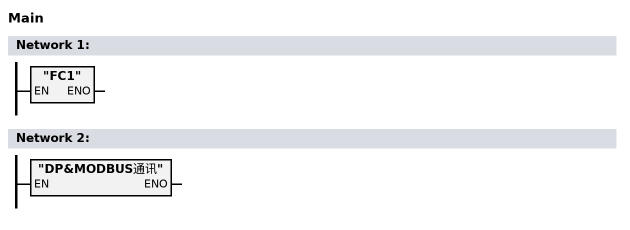
   RUNG wire#powerrail
      "FC1"()
   END_RUNG
   // the same network as SCL:
   "FC1"();
END_REGION

REGION Network 2
   RUNG wire#powerrail
      "DP&MODBUS通讯"()
   END_RUNG
   // the same network as SCL:
   "DP&MODBUS通讯"();
END_REGION
END_ORGANIZATION_BLOCK

// ===== PLC "2#GZY"  CPU 1511-1 PN =====

VAR_GLOBAL   // PLC tag table "默认变量表"
   "Clock_Byte" AT %MB0 : Byte;
   "Clock_10Hz" AT %M0.0 : Bool;
   "Clock_5Hz" AT %M0.1 : Bool;
   "Clock_2.5Hz" AT %M0.2 : Bool;
   "Clock_2Hz" AT %M0.3 : Bool;
   "Clock_1.25Hz" AT %M0.4 : Bool;
   "Clock_1Hz" AT %M0.5 : Bool;
   "Clock_0.625Hz" AT %M0.6 : Bool;
   "Clock_0.5Hz" AT %M0.7 : Bool;
   "2#干燥窑主机远程" AT %I0.0 : Bool;
   "2#干燥窑主机变频备妥" AT %I0.1 : Bool;
   "2#干燥窑主机散热风机运行" AT %I0.2 : Bool;
   "2#干燥窑变频运行" AT %I0.3 : Bool;
   "2#干燥窑变频故障" AT %I0.4 : Bool;
   "2#干燥窑稀油中控" AT %I1.0 : Bool;
   "2#干燥窑稀油1#泵运行" AT %I1.1 : Bool;
   "2#干燥窑稀油2#泵运行" AT %I1.2 : Bool;
   "2#干燥窑稀油油差下限" AT %I1.3 : Bool;
   "2#干燥窑稀油油位上限" AT %I1.4 : Bool;
   "2#干燥窑稀油油位下限" AT %I1.5 : Bool;
   "2#干燥窑稀油1#泵故障" AT %I1.6 : Bool;
   "2#干燥窑稀油2#泵故障" AT %I1.7 : Bool;
   "2#干燥窑挡轮备妥" AT %I2.0 : Bool;
   "2#干燥窑挡轮1#泵运行" AT %I2.1 : Bool;
   "2#干燥窑挡轮2#泵运行" AT %I2.2 : Bool;
   "2#干燥窑挡轮溢流阀运行" AT %I2.3 : Bool;
   "2#干燥窑挡轮行程过低" AT %I2.4 : Bool;
   "2#干燥窑挡轮故障" AT %I2.5 : Bool;
   "I3_0" AT %I3.0 : Bool;
   "I3_1" AT %I3.1 : Bool;
   "I3_2" AT %I3.2 : Bool;
   "湿矿转2#干燥窑皮中控  (3#皮带)" AT %I3.3 : Bool;
   "湿矿转2#干燥窑皮运行  (3#皮带)" AT %I3.4 : Bool;
   "湿矿转2#干燥窑皮故障  (3#皮带)" AT %I3.5 : Bool;
   "I4_0" AT %I4.0 : Bool;
   "I4_1" AT %I4.1 : Bool;
   "I4_2" AT %I4.2 : Bool;
   "I4_3" AT %I4.3 : Bool;
   "I4_4" AT %I4.4 : Bool;
   "I4_5" AT %I4.5 : Bool;
   "I5_0" AT %I5.0 : Bool;
   "I5_1" AT %I5.1 : Bool;
   "I5_2" AT %I5.2 : Bool;
   "I5_3" AT %I5.3 : Bool;
   "I5_4" AT %I5.4 : Bool;
   "I5_5" AT %I5.5 : Bool;
   "定量给煤机中控" AT %I6.3 : Bool;
   "定量给煤机运行" AT %I6.4 : Bool;
   "定量给煤机故障" AT %I6.5 : Bool;
   "定量给煤机流量脉冲" AT %I6.6 : Bool;
   "煤粉仓收尘风机中控" AT %I7.0 : Bool;
   "煤粉仓收尘风机运行" AT %I7.1 : Bool;
   "煤粉仓收尘风机故障" AT %I7.2 : Bool;
   "2#干燥窑一次风机中控" AT %I8.0 : Bool;
   "2#干燥窑一次风机运行" AT %I8.1 : Bool;
   "2#干燥窑一次风机故障" AT %I8.2 : Bool;
   "2#干燥窑二次风机中控" AT %I8.3 : Bool;
   "2#干燥窑二次风机运行" AT %I8.4 : Bool;
   "2#干燥窑二次风机故障" AT %I8.5 : Bool;
   "I9_0" AT %I9.0 : Bool;
   "I9_1" AT %I9.1 : Bool;
   "I9_2" AT %I9.2 : Bool;
   "I9_3" AT %I9.3 : Bool;
   "I9_4" AT %I9.4 : Bool;
   "I9_5" AT %I9.5 : Bool;
   "I10_0" AT %I10.0 : Bool;
   "I10_1" AT %I10.1 : Bool;
   "I10_2" AT %I10.2 : Bool;
   "I10_4" AT %I10.4 : Bool;
   "I10_5" AT %I10.5 : Bool;
   "I10_6" AT %I10.6 : Bool;
   "2#干燥窑转速" AT %IW256 : Int;
   "2#干燥窑电流" AT %IW258 : Int;
   "PIW260" AT %IW260 : Int;
   "2#干燥窑一次风机电流" AT %IW262 : Int;
   "2#干燥窑二次风机频率" AT %IW264 : Int;
   "2#干燥窑二次风机电流" AT %IW266 : Int;
   "PIW268" AT %IW268 : Int;
   "PIW270" AT %IW270 : Int;
   "2#干燥窑窑尾压力" AT %IW272 : Int;
   "PIW274" AT %IW274 : Int;
   "定量给煤机流量" AT %IW276 : Int;
   "烟气管道进口压力" AT %IW278 : Int;
   "2#干燥窑一次风压" AT %IW280 : Int;
   "2#干燥窑二次风压" AT %IW282 : Int;
   "煤粉仓压力" AT %IW284 : Int;
   "混合室压力" AT %IW286 : Int;
   "煤粉仓温度1(PT100)" AT %IW288 : Int;
   "煤粉仓温度2(PT100)" AT %IW290 : Int;
   "煤粉仓温度3(PT100)" AT %IW292 : Int;
   "煤粉仓温度4(PT100)" AT %IW294 : Int;
   "窑尾温度 K偶" AT %IW296 : Int;
   "烟气管道进口温度 K偶" AT %IW298 : Int;
   "燃烧室温度 4~20mA" AT %IW300 : Int;
   "混合室温度 4~20mA" AT %IW302 : Int;
   "2#窑A档轴温1" AT %ID320 : Real;
   "2#窑A档油温1" AT %ID324 : Real;
   "2#窑A档轴温2" AT %ID328 : Real;
   "2#窑A档油温2" AT %ID332 : Real;
   "2#窑A档轴温3" AT %ID336 : Real;
   "2#窑A档油温3" AT %ID340 : Real;
   "2#窑A档轴温4" AT %ID344 : Real;
   "2#窑A档油温4" AT %ID348 : Real;
   "2#窑B档轴温1" AT %ID352 : Real;
   "2#窑B档油温1" AT %ID356 : Real;
   "2#窑B档轴温2" AT %ID360 : Real;
   "2#窑B档油温2" AT %ID364 : Real;
   "2#窑B档轴温3" AT %ID368 : Real;
   "2#窑B档油温3" AT %ID372 : Real;
   "2#窑B档轴温4" AT %ID376 : Real;
   "2#窑B档油温4" AT %ID380 : Real;
   "2#窑主电机A相绕组温度" AT %ID384 : Real;
   "干燥窑主传动合闸" AT %Q0.0 : Bool;
   "干燥窑主传动分闸" AT %Q0.1 : Bool;
   "干燥窑主传动变频启动" AT %Q0.2 : Bool;
   "干燥窑主传稀油站启动" AT %Q0.3 : Bool;
   "湿矿转2#干燥窑皮带启动  (3#皮带)" AT %Q0.4 : Bool;
   "Q0_5" AT %Q0.5 : Bool;
   "Q0_6" AT %Q0.6 : Bool;
   "Q0_7" AT %Q0.7 : Bool;
   "Q1_0" AT %Q1.0 : Bool;
   "定量给煤机启动" AT %Q1.2 : Bool;
   "煤粉仓收尘风机启动" AT %Q1.3 : Bool;
   "Q1_4" AT %Q1.4 : Bool;
   "Q1_5" AT %Q1.5 : Bool;
   "干燥窑挡轮油站启动" AT %Q1.6 : Bool;
   "2#干燥窑一次风机启动" AT %Q2.0 : Bool;
   "2#干燥窑二次风机启动" AT %Q2.1 : Bool;
   "Q2_2" AT %Q2.2 : Bool;
   "Q2_3" AT %Q2.3 : Bool;
   "Tag_8" AT %QB4 : Byte;
   "2#干燥窑转速给定" AT %QW256 : Int;
   "定量给煤机流量给定" AT %QW258 : Int;
   "PQW264" AT %QW264 : Int;
   "2#干燥窑二次风机频率给定" AT %QW266 : Int;
   "PQW268" AT %QW268 : Int;
   "PQW270" AT %QW270 : Int;
   "Tag_1" AT %MW4 : Word;
   "Tag_2" AT %M400.0 : Bool;
   "连锁解锁" AT %M400.2 : Bool;
   "干燥窑连锁信号" AT %M400.3 : Bool;
   "Tag_4" AT %M400.5 : Bool;
   "Tag_5" AT %MW410 : Word;
   "Tag_6" AT %MW412 : Word;
   "稀油站油压长时间低" AT %T6 : Timer;
   "稀油站启动10S" AT %T7 : Timer;
   "稀油站油差下限时间" AT %T8 : Timer;
   "Tag_3" AT %C1 : Counter;
   "Tag_7" AT %C2 : Counter;
   "2#干燥窑断路器合闸" AT %I0.5 : Bool;
   "2#干燥窑断路器分闸" AT %I0.6 : Bool;
   "2#干燥窑进料口压力" AT %IW304 : Int;
   "Tag_31" AT %T1 : Timer;
   "Tag_33" AT %T2 : Timer;
   "Q1_1" AT %Q1.1 : Bool;
   "System_Byte" AT %MB1 : Byte;
   "FirstScan" AT %M1.0 : Bool;
   "DiagStatusUpdate" AT %M1.1 : Bool;
   "AlwaysTRUE" AT %M1.2 : Bool;
   "AlwaysFALSE" AT %M1.3 : Bool;
   "2#窑主电机B相绕组温度" AT %ID388 : Real;
   "2#窑主电机C相绕组温度" AT %ID392 : Real;
   "2#窑主电机前轴承温度" AT %ID396 : Real;
   "2#窑主电机后轴承温度" AT %ID400 : Real;
   "I0_7" AT %I0.7 : Bool;
   "I2_6" AT %I2.6 : Bool;
   "I2_7" AT %I2.7 : Bool;
   "I3_6" AT %I3.6 : Bool;
   "I3_7" AT %I3.7 : Bool;
   "I4_6" AT %I4.6 : Bool;
   "I4_7" AT %I4.7 : Bool;
   "I5_6" AT %I5.6 : Bool;
   "I5_7" AT %I5.7 : Bool;
   "I6_0" AT %I6.0 : Bool;
   "I6_1" AT %I6.1 : Bool;
   "I6_2" AT %I6.2 : Bool;
   "I6_7" AT %I6.7 : Bool;
   "I7_3" AT %I7.3 : Bool;
   "I7_4" AT %I7.4 : Bool;
   "I7_5" AT %I7.5 : Bool;
   "I7_6" AT %I7.6 : Bool;
   "I7_7" AT %I7.7 : Bool;
   "I8_6" AT %I8.6 : Bool;
   "I8_7" AT %I8.7 : Bool;
   "I9_6" AT %I9.6 : Bool;
   "I9_7" AT %I9.7 : Bool;
   "I10_3" AT %I10.3 : Bool;
   "I10_7" AT %I10.7 : Bool;
   "I11_0" AT %I11.0 : Bool;
   "I11_1" AT %I11.1 : Bool;
   "I11_2" AT %I11.2 : Bool;
   "I11_3" AT %I11.3 : Bool;
   "I11_4" AT %I11.4 : Bool;
   "I11_5" AT %I11.5 : Bool;
   "I11_6" AT %I11.6 : Bool;
   "I11_7" AT %I11.7 : Bool;
   "Q1_7" AT %Q1.7 : Bool;
   "Q2_4" AT %Q2.4 : Bool;
   "Q2_5" AT %Q2.5 : Bool;
   "Q2_6" AT %Q2.6 : Bool;
   "Q2_7" AT %Q2.7 : Bool;
   "Q3_0" AT %Q3.0 : Bool;
   "Q3_1" AT %Q3.1 : Bool;
   "Q3_2" AT %Q3.2 : Bool;
   "Q3_3" AT %Q3.3 : Bool;
   "Q3_4" AT %Q3.4 : Bool;
   "Q3_5" AT %Q3.5 : Bool;
   "Q3_6" AT %Q3.6 : Bool;
   "Q3_7" AT %Q3.7 : Bool;
   "2#给煤机出料口负压" AT %IW306 : Int;
   "PIW308" AT %IW308 : Int;
   "PIW310" AT %IW310 : Int;
   "PIW312" AT %IW312 : Int;
   "PIW314" AT %IW314 : Int;
   "PIW316" AT %IW316 : Int;
   "PIW318" AT %IW318 : Int;
   "PQW260" AT %QW260 : Int;
   "PQW262" AT %QW262 : Int;
   "2#干燥窑煤粉仓称重" AT %ID440 : Real;
   "Tag_9" AT %T10 : Timer;
END_VAR

DATA_BLOCK "驱动"   // DB1
{ S7_Optimized_Access := 'FALSE' }
VERSION : 0.1
   VAR
      "2#二次风机启动" : Bool;
      "2#二次风机停止" : Bool;
      "2#干燥窑主机合闸" : Bool;
      "2#干燥窑主机分闸" : Bool;
      STAT4 : Bool;
      STAT5 : Bool;
      "2#干燥窑主机启动" : Bool;
      "2#干燥窑主机停止" : Bool;
      STAT8 : Bool;
      STAT9 : Bool;
      STAT10 : Bool;
      STAT11 : Bool;
      "gzy进窑2#皮带启动3#皮带" : Bool;
      "gzy进窑2#皮带停止3#皮带" : Bool;
      STAT14 : Bool;
      STAT15 : Bool;
      STAT16 : Bool;
      STAT17 : Bool;
      STAT18 : Bool;
      STAT19 : Bool;
      STAT20 : Bool;
      STAT21 : Bool;
      STAT22 : Bool;
      STAT23 : Bool;
      STAT24 : Bool;
      STAT25 : Bool;
      STAT26 : Bool;
      STAT27 : Bool;
      "2#一次风机启动" : Bool;
      "2#一次风机停止" : Bool;
      STAT30 : Bool;
      STAT31 : Bool;
      STAT32 : Bool;
      STAT33 : Bool;
      STAT34 : Bool;
      STAT35 : Bool;
      STAT36 : Bool;
      STAT37 : Bool;
      STAT38 : Bool;
      STAT39 : Bool;
      "2#干燥窑煤粉收尘风机启动" : Bool;
      "2#干燥窑煤粉收尘风机停止" : Bool;
      "2#干燥窑锁风给煤机启动" : Bool;
      "2#干燥窑锁风给煤机停止" : Bool;
      "2#干燥窑锁风给煤机分割轮启动" : Bool;
      "2#干燥窑锁风给煤机分割轮停止" : Bool;
      STAT46 : Bool;
      STAT47 : Bool;
      STAT48 : Bool;
      STAT49 : Bool;
      STAT50 : Bool;
      STAT51 : Bool;
      STAT52 : Bool;
      STAT53 : Bool;
      STAT54 : Bool;
      STAT55 : Bool;
      STAT56 : Bool;
      "2#干燥窑联锁解锁" : Bool;
      STAT58 : Bool;
      STAT59 : Bool;
      STAT60 : Bool;
      "2#干燥窑定量给煤机班累计清零" : Bool;
      "2#干燥窑定量给煤机日累计清零" : Bool;
      "2#干燥窑定量给煤机总累计清零" : Bool;
      STAT64 : Bool;
      STAT65 : Bool;
      "2#干燥窑稀油站启动" : Bool;
      "2#干燥窑稀油站停止" : Bool;
      "2#干燥窑挡轮油站启动" : Bool;
      "2#干燥窑挡轮油站停止" : Bool;
      STAT66 : Bool;
      STAT67 : Bool;
   END_VAR
BEGIN
END_DATA_BLOCK

DATA_BLOCK "模拟量"   // DB2
{ S7_Optimized_Access := 'FALSE' }
VERSION : 0.1
   VAR
      STAT0 : Int;
      STAT1 : Int;
      STAT2 : Int;
      STAT3 : Int;
      STAT4 : Int;
      STAT5 : Int;
      STAT6 : Int;
      STAT7 : Int;
      STAT8 : Int;
      STAT9 : Real;
      STAT10 : Real;
      STAT11 : Real;
      STAT12 : Real;
      STAT13 : Real;
      STAT14 : Real;
      STAT15 : Real;
      STAT16 : Real;
      STAT17 : Real;
      STAT18 : Real;
      STAT19 : Real;
      STAT20 : Real;
      STAT21 : Real;
      STAT22 : Real;
      STAT23 : Real;
      STAT24 : Real;
      STAT25 : Real;
      STAT26 : Real;
      STAT27 : Real;
      STAT28 : Real;
      STAT29 : Real;
      STAT30 : Real;
      STAT31 : Real;
      STAT32 : Real;
      STAT33 : Real;
      STAT34 : Real;
      STAT35 : Real;
      STAT36 : Real;
      STAT37 : Real;
      STAT38 : Real;
      STAT39 : Real;
      STAT40 : Real;
      STAT41 : Real;
      STAT42 : Real;
      STAT43 : Real;
      STAT44 : Real;
      STAT45 : Real;
      STAT46 : Real;
      STAT47 : Real;
      STAT48 : Real;
      STAT49 : Real;
      STAT50 : Real;
      STAT51 : Real;
      STAT52 : Real;
      STAT53 : Real;
      STAT54 : Real;
      STAT55 : Real;
      STAT56 : Real;
      STAT57 : Real;
      STAT58 : Real;
      STAT59 : Real;
      STAT60 : Real;
      STAT61 : Real;
      STAT62 : Real;
      STAT63 : Real;
      STAT64 : Real;
      STAT65 : Real;
      STAT66 : Real;
      STAT67 : Real;
      STAT68 : Real;
      STAT69 : Real;
      STAT70 : Real;
      STAT71 : Real;
      STAT72 : Real;
      STAT73 : Real;
      STAT74 : Real;
      STAT75 : Real;
      STAT76 : Real;
      STAT77 : Real;
      STAT78 : Real;
      STAT79 : Real;
      STAT80 : Real;
      STAT81 : Real;
   END_VAR
BEGIN
END_DATA_BLOCK

DATA_BLOCK "给煤机班累计DB块"   // DB3
{ S7_Optimized_Access := 'FALSE' }
VERSION : 0.0
// stored: InstanceOfName 累计功能块
"累计功能块"
BEGIN
END_DATA_BLOCK

DATA_BLOCK "给煤机日累计DB块"   // DB4
{ S7_Optimized_Access := 'FALSE' }
VERSION : 0.0
// stored: InstanceOfName 累计功能块
"累计功能块"
BEGIN
END_DATA_BLOCK

DATA_BLOCK "给煤机总累计DB块"   // DB5
{ S7_Optimized_Access := 'FALSE' }
VERSION : 0.0
// stored: InstanceOfName 累计功能块
"累计功能块"
BEGIN
END_DATA_BLOCK

DATA_BLOCK "DB6_皮带秤粘料"   // DB6
{ S7_Optimized_Access := 'FALSE' }
VERSION : 0.1
   VAR
      干燥窑定量给煤机给定反馈差值 : Real;
      干燥窑定量给煤机给定反馈差值绝对值 : Real;
      real3 : Real;
      real4 : Real;
      real5 : Real;
      real6 : Real;
      real7 : Real;
      real8 : Real;
      real9 : Real;
      real10 : Real;
      real11 : Real;
      real12 : Real;
      real13 : Real;
      real14 : Real;
      real15 : Real;
      real16 : Real;
      real17 : Real;
      real18 : Real;
      real19 : Real;
      real20 : Real;
      干燥窑定量给煤机粘料报警 : Bool;
      bool2 : Bool;
      bool3 : Bool;
      bool4 : Bool;
      bool5 : Bool;
      bool6 : Bool;
      bool7 : Bool;
      bool8 : Bool;
      bool9 : Bool;
      bool10 : Bool;
      bool11 : Bool;
      bool12 : Bool;
      bool13 : Bool;
      bool14 : Bool;
      bool15 : Bool;
      bool16 : Bool;
      bool17 : Bool;
      bool18 : Bool;
      bool19 : Bool;
      bool20 : Bool;
      bool21 : Bool;
   END_VAR
BEGIN
END_DATA_BLOCK

DATA_BLOCK "累计功能块2_DB"   // DB7
{ S7_Optimized_Access := 'FALSE' }
VERSION : 0.1
// stored: InstanceOfName 累计功能块2
"累计功能块2"
BEGIN
END_DATA_BLOCK

DATA_BLOCK "通讯仪表数据"   // DB20
{ S7_Optimized_Access := 'FALSE' }
VERSION : 0.1
   VAR
      STAT0 : Int;
      "1#窑A档油温1" : Real := 33.4;
      "1#窑A档油温2" : Real := 33.0;
      "1#窑A档油温3" : Real := 34.3;
      "1#窑A档油温4" : Real := 34.0;
      "1#窑A档轴温1" : Real := 33.6;
      "1#窑A档轴温2" : Real := 33.4;
      "1#窑A档轴温3" : Real := 33.6;
      "1#窑A档轴温4" : Real := 34.5;
      "1#窑B档油温1" : Real := 34.3;
      "1#窑B档油温2" : Real := 34.5;
      "1#窑B档油温3" : Real := 35.0;
      "1#窑B档油温4" : Real := 36.1;
      "1#窑B档轴温1" : Real := 34.9;
      "1#窑B档轴温2" : Real := 36.4;
      "1#窑B档轴温3" : Real := 34.9;
      "1#窑B档轴温4" : Real := 36.2;
      "1#窑主电机A相绕组温度" : Real := 62.7;
      "1#窑主电机B相绕组温度" : Real := 63.4;
      "1#窑主电机C相绕组温度" : Real := 62.0;
      "1#窑主电机前轴承温度" : Real := 45.0;
      "1#窑主电机后轴承温度" : Real := 41.8;
      STAT22 : Real;
      STAT23 : Real;
      STAT24 : Real;
      STAT25 : Real;
      STAT26 : Real;
      STAT27 : Real;
      STAT28 : Real;
      STAT29 : Real;
      STAT30 : Real;
      STAT31 : Real;
      STAT32 : Real;
      "1#干燥窑煤粉仓称重" : Real := 11.52;   // 1#干燥窑煤粉仓称重
      STAT34 : Real;
   END_VAR
BEGIN
END_DATA_BLOCK

DATA_BLOCK "模拟量数据"   // DB21
{ S7_Optimized_Access := 'FALSE' }
VERSION : 0.1
   VAR
      "2#干燥窑主电机转速" : Real := 798.1337;
      "2#干燥窑主电机电流" : Real := 254.8892;
      STAT2 : Real;
      "2#干燥窑一次风机运行电流" : Real;
      "2#二次风机运行频率" : Real := 33.52141;
      "2#二次风机运行电流" : Real := 98.98177;
      STAT6 : Real;
      STAT7 : Real;
      "2#干燥窑窑尾烟气管道压力" : Real := -500.0;
      STAT9 : Real;
      "2#干燥窑煤粉流量" : Real := 2.009259;
      "2#干燥窑进口烟气管道压力" : Real := -1000.0;
      "2#干燥窑一次风机压力" : Real := 2973.09;
      "2#干燥窑二次风机压力" : Real := 1742.188;
      "2#干燥窑煤粉仓压力" : Real := 4.340332;
      "2#干燥窑燃烧室压力" : Real := -913.6285;
      "2#干燥窑煤粉仓温度1" : Real := 34.20139;
      "2#干燥窑煤粉仓温度2" : Real := 33.85416;
      "2#干燥窑煤粉仓温度3" : Real := 33.44907;
      "2#干燥窑煤粉仓温度4" : Real := 32.55209;
      "2#干燥窑窑尾罩温度" : Real := 136.169;
      "2#干燥窑进口烟气管道温度" : Real := 201.6204;
      "2#干燥窑燃烧室温度" : Real := 877.3149;
      "2#干燥窑混合室温度" : Real := 512.7025;
      "2#干燥窑主电机转速给定" : Real := 800.0;
      "2#干燥窑煤粉仓流量给定" : Real := 2.0;
      STAT26 : Real;
      STAT27 : Real;
      STAT28 : Real;
      "2#二次风机频率给定" : Real := 33.0;
      STAT30 : Real;
      STAT31 : Real;
      "2#干燥窑定量给煤机班累计" : Real := 0.0322427;
      "2#干燥窑定量给煤机日累计" : Real := 312.7758;
      "2#干燥窑定量给煤机总累计" : Real := 312.7776;
      STAT35 : Real;
      STAT36 : Real;
   END_VAR
BEGIN
END_DATA_BLOCK

DATA_BLOCK "窑联锁数据DB块"   // DB23
{ S7_Optimized_Access := 'FALSE' }
VERSION : 0.1
   VAR
      STAT0 : Bool := TRUE;
      STAT1 : Bool;
      STAT2 : Bool;
      STAT3 : Bool;
      STAT4 : Bool;
      STAT5 : Bool;
      STAT6 : Bool;
      STAT7 : Bool;
      STAT8 : Bool := TRUE;
      STAT9 : Bool;
      STAT10 : Bool;
      STAT11 : Bool;
      STAT12 : Bool;
      STAT13 : Bool;
      STAT14 : Bool;
      STAT15 : Bool;
      STAT16 : Bool;
      STAT17 : Bool;
      STAT18 : Word;
   END_VAR
BEGIN
END_DATA_BLOCK

DATA_BLOCK "DB26"   // DB26
{ S7_Optimized_Access := 'FALSE' }
VERSION : 0.1
   VAR
      STAT0 : Bool;
      STAT1 : Bool;
      STAT2 : Bool;
      STAT3 : Bool;
      STAT4 : Bool;
      STAT5 : Bool;
      STAT6 : Bool;
      STAT7 : Bool;
      STAT8 : Word := WORD#16#0002;
      STAT9 : Word;
      STAT10 : Word;
   END_VAR
BEGIN
END_DATA_BLOCK

DATA_BLOCK "FB40_DATA_ALARM_DB"   // DB40
{ S7_Optimized_Access := 'FALSE' }
VERSION : 0.1
// stored: InstanceOfName FB40_DATA_ALARM
"FB40_DATA_ALARM"
BEGIN
END_DATA_BLOCK

FUNCTION_BLOCK "累计功能块"   // FB10, STL
{ S7_Optimized_Access := 'FALSE' }
VERSION : 0.1
   VAR_INPUT
      IN0 : Real;
      IN1 : Bool;
   END_VAR
   VAR_OUTPUT
      OUT2 : Real;
   END_VAR
   VAR
      STAT3 : Real;
      STAT4 : Real;
      STAT5 : Real;
   END_VAR
BEGIN

REGION Network 1
         A(;
         A(;
         A(;
         L     #IN0;
         L     3600.0;
         /R;
         T     #STAT3;
         AN    OV;
         SAVE;
         CLR;
         A     BR;
         );
         JNB   M001;
         L     #STAT3;
         L     10.0;
         /R;
         T     #STAT4;
         AN    OV;
         SAVE;
         CLR;
   M001: A     BR;
         );
         JNB   M002;
         L     #STAT4;
         L     #STAT5;
         +R;
         T     #STAT5;
         AN    OV;
         SAVE;
         CLR;
   M002: A     BR;
         );
         JNB   M003;
         L     #STAT5;
         T     #OUT2;
   M003: NOP   0;
END_REGION

REGION Network 2
         A     #IN1;
         =     %L0.0;
         A     %L0.0;
         JNB   M004;
         L     0.0;
         T     #STAT3;
   M004: NOP   0;
         A     %L0.0;
         JNB   M005;
         L     0.0;
         T     #STAT4;
   M005: NOP   0;
         A     %L0.0;
         JNB   M006;
         L     0.0;
         T     #STAT5;
   M006: NOP   0;
END_REGION

REGION Network 3
         SET;
         SAVE;
END_REGION
END_FUNCTION_BLOCK

FUNCTION_BLOCK "FB40_DATA_ALARM"   // FB40, LAD
{ S7_Optimized_Access := 'FALSE' }
VERSION : 0.1
   VAR
      "2#干燥窑转速" : "FB330_DATA_ALARM";
      "2#干燥窑电流" : "FB330_DATA_ALARM";
      PIW260 : "FB330_DATA_ALARM";
      "2#干燥窑一次风机电流" : "FB330_DATA_ALARM";
      "2#干燥窑二次风机频率" : "FB330_DATA_ALARM";
      "2#干燥窑二次风机电流" : "FB330_DATA_ALARM";
      PIW268 : "FB330_DATA_ALARM";
      PIW270 : "FB330_DATA_ALARM";
      "2#干燥窑窑尾压力" : "FB330_DATA_ALARM";
      PIW274 : "FB330_DATA_ALARM";
      定量给煤机流量 : "FB330_DATA_ALARM";
      烟气管道进口压力 : "FB330_DATA_ALARM";
      "2#干燥窑一次风压" : "FB330_DATA_ALARM";
      "2#干燥窑二次风压" : "FB330_DATA_ALARM";
      煤粉仓压力 : "FB330_DATA_ALARM";
      混合室压力 : "FB330_DATA_ALARM";
      "煤粉仓温度1(PT100)" : "FB330_DATA_ALARM";
      "煤粉仓温度2(PT100)" : "FB330_DATA_ALARM";
      "煤粉仓温度3(PT100)" : "FB330_DATA_ALARM";
      "煤粉仓温度4(PT100)" : "FB330_DATA_ALARM";
      "窑尾温度 K偶" : "FB330_DATA_ALARM";
      "烟气管道进口温度 K偶" : "FB330_DATA_ALARM";
      "燃烧室温度 4~20mA" : "FB330_DATA_ALARM";
      "混合室温度 4~20mA" : "FB330_DATA_ALARM";
      "2#干燥窑进料口压力" : "FB330_DATA_ALARM";
      "2#给煤机出料口负压" : "FB330_DATA_ALARM";
      PIW308 : "FB330_DATA_ALARM";
      PIW310 : "FB330_DATA_ALARM";
      PIW312 : "FB330_DATA_ALARM";
      PIW314 : "FB330_DATA_ALARM";
      PIW316 : "FB330_DATA_ALARM";
      PIW318 : "FB330_DATA_ALARM";
      "2#窑A档轴温1" : "FB330_DATA_ALARM";
      "2#窑A档油温1" : "FB330_DATA_ALARM";
      "2#窑A档轴温2" : "FB330_DATA_ALARM";
      "2#窑A档油温2" : "FB330_DATA_ALARM";
      "2#窑A档轴温3" : "FB330_DATA_ALARM";
      "2#窑A档油温3" : "FB330_DATA_ALARM";
      "2#窑A档轴温4" : "FB330_DATA_ALARM";
      "2#窑A档油温4" : "FB330_DATA_ALARM";
      "2#窑B档轴温1" : "FB330_DATA_ALARM";
      "2#窑B档油温1" : "FB330_DATA_ALARM";
      "2#窑B档轴温2" : "FB330_DATA_ALARM";
      "2#窑B档油温2" : "FB330_DATA_ALARM";
      "2#窑B档轴温3" : "FB330_DATA_ALARM";
      "2#窑B档油温3" : "FB330_DATA_ALARM";
      "2#窑B档轴温4" : "FB330_DATA_ALARM";
      "2#窑B档油温4" : "FB330_DATA_ALARM";
      "2#窑主电机A相绕组温度" : "FB330_DATA_ALARM";
      "2#窑主电机B相绕组温度" : "FB330_DATA_ALARM";
      "2#窑主电机C相绕组温度" : "FB330_DATA_ALARM";
      "2#窑主电机前轴承温度" : "FB330_DATA_ALARM";
      "2#窑主电机后轴承温度" : "FB330_DATA_ALARM";
      PID404 : "FB330_DATA_ALARM";
      PID408 : "FB330_DATA_ALARM";
      PID412 : "FB330_DATA_ALARM";
      "2#干燥窑煤粉仓称重" : "FB330_DATA_ALARM";
      STATIC1 : "FB330_DATA_ALARM";
      STATIC2 : "FB330_DATA_ALARM";
      STATIC3 : "FB330_DATA_ALARM";
   END_VAR
   VAR_TEMP
      TEMP1 : Real;
   END_VAR
BEGIN

REGION Network 1
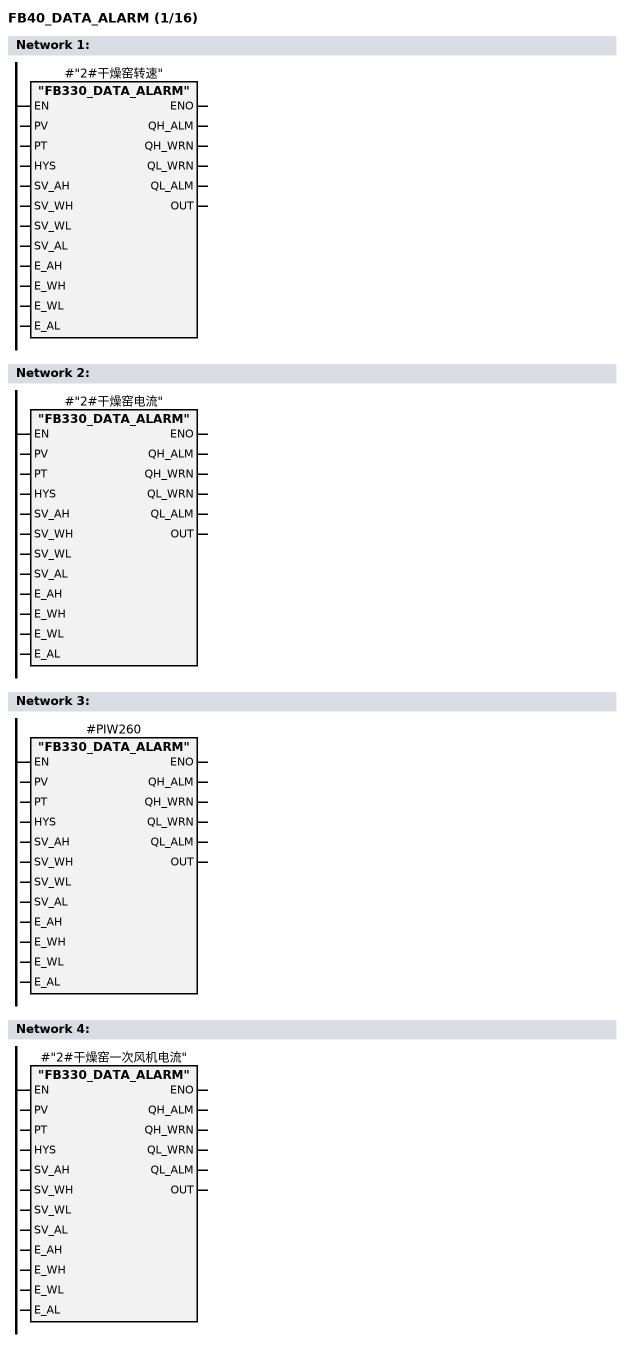
   RUNG wire#powerrail
      #"2#干燥窑转速"(PV :=, PT :=, HYS :=, SV_AH :=, SV_WH :=, SV_WL :=, SV_AL :=, E_AH :=, E_WH :=, E_WL :=, E_AL :=, QH_ALM =>, QH_WRN =>, QL_WRN =>, QL_ALM =>, OUT =>)
   END_RUNG
   // the same network as SCL:
   #"2#干燥窑转速"();   // "FB330_DATA_ALARM"
END_REGION

REGION Network 2
   RUNG wire#powerrail
      #"2#干燥窑电流"(PV :=, PT :=, HYS :=, SV_AH :=, SV_WH :=, SV_WL :=, SV_AL :=, E_AH :=, E_WH :=, E_WL :=, E_AL :=, QH_ALM =>, QH_WRN =>, QL_WRN =>, QL_ALM =>, OUT =>)
   END_RUNG
   // the same network as SCL:
   #"2#干燥窑电流"();   // "FB330_DATA_ALARM"
END_REGION

REGION Network 3
   RUNG wire#powerrail
      #PIW260(PV :=, PT :=, HYS :=, SV_AH :=, SV_WH :=, SV_WL :=, SV_AL :=, E_AH :=, E_WH :=, E_WL :=, E_AL :=, QH_ALM =>, QH_WRN =>, QL_WRN =>, QL_ALM =>, OUT =>)
   END_RUNG
   // the same network as SCL:
   #PIW260();   // "FB330_DATA_ALARM"
END_REGION

REGION Network 4
   RUNG wire#powerrail
      #"2#干燥窑一次风机电流"(PV :=, PT :=, HYS :=, SV_AH :=, SV_WH :=, SV_WL :=, SV_AL :=, E_AH :=, E_WH :=, E_WL :=, E_AL :=, QH_ALM =>, QH_WRN =>, QL_WRN =>, QL_ALM =>, OUT =>)
   END_RUNG
   // the same network as SCL:
   #"2#干燥窑一次风机电流"();   // "FB330_DATA_ALARM"
END_REGION

REGION Network 5
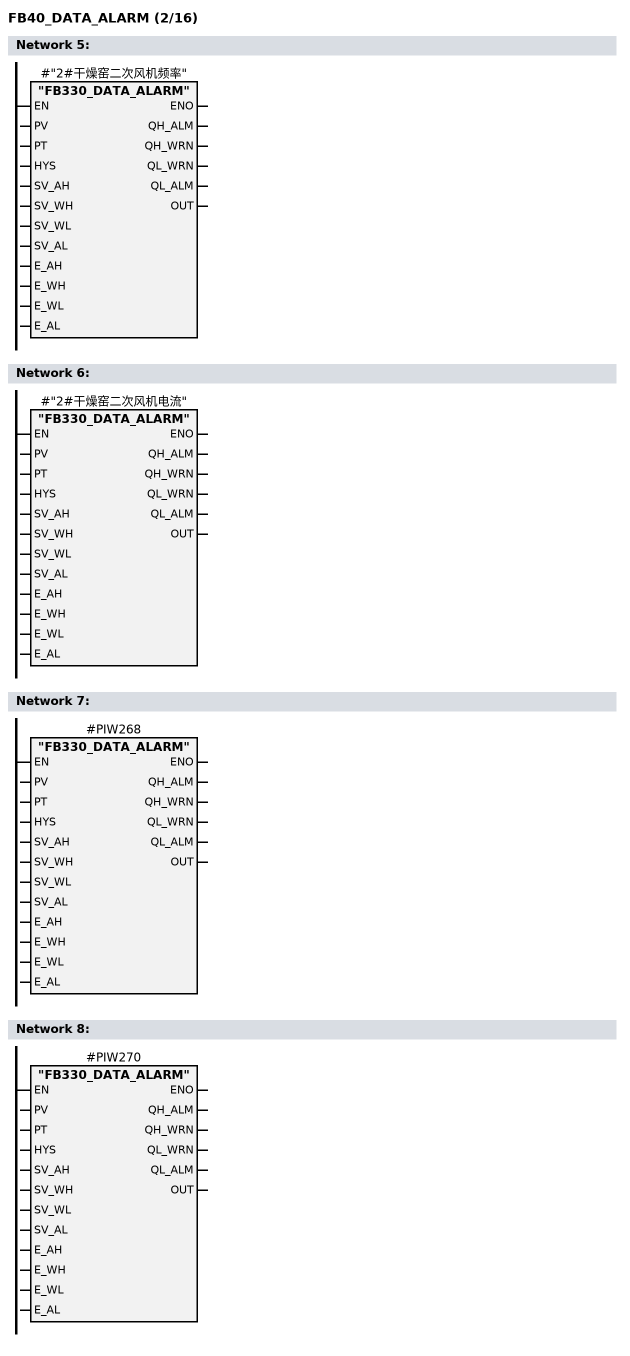
   RUNG wire#powerrail
      #"2#干燥窑二次风机频率"(PV :=, PT :=, HYS :=, SV_AH :=, SV_WH :=, SV_WL :=, SV_AL :=, E_AH :=, E_WH :=, E_WL :=, E_AL :=, QH_ALM =>, QH_WRN =>, QL_WRN =>, QL_ALM =>, OUT =>)
   END_RUNG
   // the same network as SCL:
   #"2#干燥窑二次风机频率"();   // "FB330_DATA_ALARM"
END_REGION

REGION Network 6
   RUNG wire#powerrail
      #"2#干燥窑二次风机电流"(PV :=, PT :=, HYS :=, SV_AH :=, SV_WH :=, SV_WL :=, SV_AL :=, E_AH :=, E_WH :=, E_WL :=, E_AL :=, QH_ALM =>, QH_WRN =>, QL_WRN =>, QL_ALM =>, OUT =>)
   END_RUNG
   // the same network as SCL:
   #"2#干燥窑二次风机电流"();   // "FB330_DATA_ALARM"
END_REGION

REGION Network 7
   RUNG wire#powerrail
      #PIW268(PV :=, PT :=, HYS :=, SV_AH :=, SV_WH :=, SV_WL :=, SV_AL :=, E_AH :=, E_WH :=, E_WL :=, E_AL :=, QH_ALM =>, QH_WRN =>, QL_WRN =>, QL_ALM =>, OUT =>)
   END_RUNG
   // the same network as SCL:
   #PIW268();   // "FB330_DATA_ALARM"
END_REGION

REGION Network 8
   RUNG wire#powerrail
      #PIW270(PV :=, PT :=, HYS :=, SV_AH :=, SV_WH :=, SV_WL :=, SV_AL :=, E_AH :=, E_WH :=, E_WL :=, E_AL :=, QH_ALM =>, QH_WRN =>, QL_WRN =>, QL_ALM =>, OUT =>)
   END_RUNG
   // the same network as SCL:
   #PIW270();   // "FB330_DATA_ALARM"
END_REGION

REGION Network 9
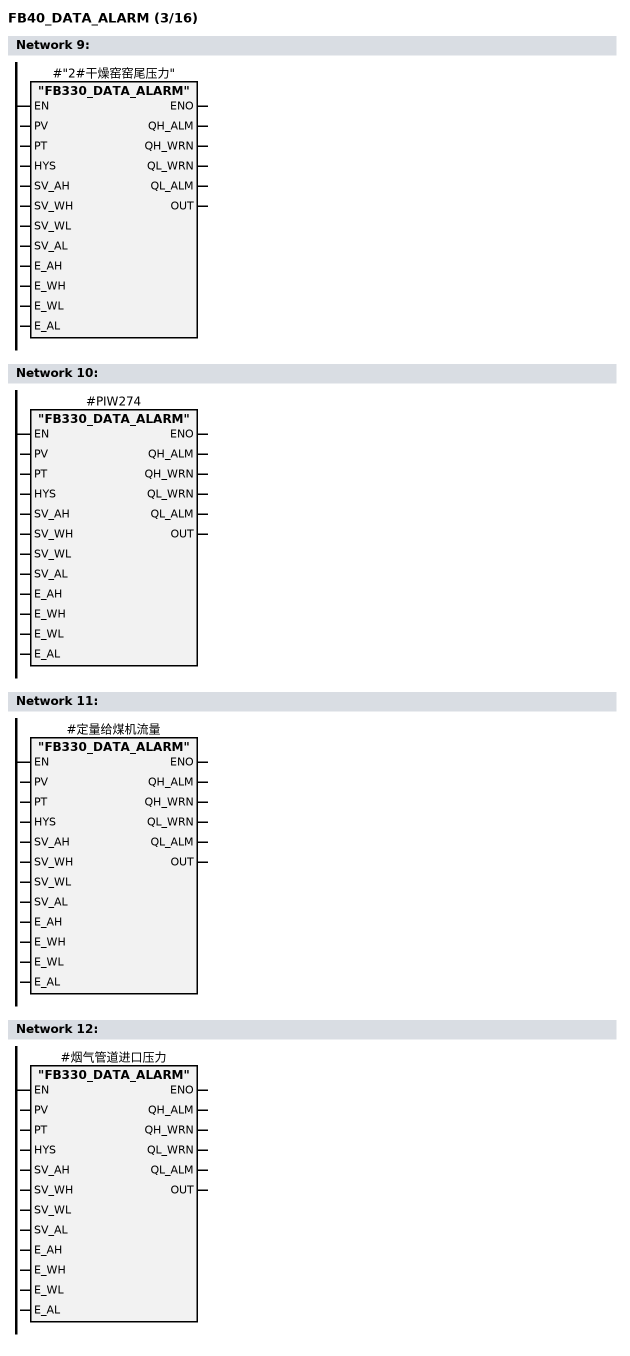
   RUNG wire#powerrail
      #"2#干燥窑窑尾压力"(PV :=, PT :=, HYS :=, SV_AH :=, SV_WH :=, SV_WL :=, SV_AL :=, E_AH :=, E_WH :=, E_WL :=, E_AL :=, QH_ALM =>, QH_WRN =>, QL_WRN =>, QL_ALM =>, OUT =>)
   END_RUNG
   // the same network as SCL:
   #"2#干燥窑窑尾压力"();   // "FB330_DATA_ALARM"
END_REGION

REGION Network 10
   RUNG wire#powerrail
      #PIW274(PV :=, PT :=, HYS :=, SV_AH :=, SV_WH :=, SV_WL :=, SV_AL :=, E_AH :=, E_WH :=, E_WL :=, E_AL :=, QH_ALM =>, QH_WRN =>, QL_WRN =>, QL_ALM =>, OUT =>)
   END_RUNG
   // the same network as SCL:
   #PIW274();   // "FB330_DATA_ALARM"
END_REGION

REGION Network 11
   RUNG wire#powerrail
      #定量给煤机流量(PV :=, PT :=, HYS :=, SV_AH :=, SV_WH :=, SV_WL :=, SV_AL :=, E_AH :=, E_WH :=, E_WL :=, E_AL :=, QH_ALM =>, QH_WRN =>, QL_WRN =>, QL_ALM =>, OUT =>)
   END_RUNG
   // the same network as SCL:
   #定量给煤机流量();   // "FB330_DATA_ALARM"
END_REGION

REGION Network 12
   RUNG wire#powerrail
      #烟气管道进口压力(PV :=, PT :=, HYS :=, SV_AH :=, SV_WH :=, SV_WL :=, SV_AL :=, E_AH :=, E_WH :=, E_WL :=, E_AL :=, QH_ALM =>, QH_WRN =>, QL_WRN =>, QL_ALM =>, OUT =>)
   END_RUNG
   // the same network as SCL:
   #烟气管道进口压力();   // "FB330_DATA_ALARM"
END_REGION

REGION Network 13